(* Logix 5000 project; controller _GigaDiscovery vendor 1 type 14 code 244 rev 35.11; software revision 35.03; part 13 of 23 *)
(* tags used below, declared in another part *)
   OS : DINT;
   Timer : TIMER[60];
   CCW_OS_Direction_1 : BOOL;
   CCW_OS_Direction_2 : BOOL;
   CROUT_Air_Compressor : UDT_CROUT;   // Compressor Command -Q18101E
   CW_OS_Direction_1 : BOOL;
   CW_OS_Direction_2 : BOOL;
   DC_Field_Pylon_Motors : UDT_CROUT;   // DC Field Pylon Motors Contactor -Q10101E -Q10103E
   Emergencies_CL0 : DINT[8];
   Emergencies_CL1 : DINT[14];
   Gate_Entry_Unlock_Selector : BOOL;   // -S30701F
   Gate_Exit_Unlock_Selector : BOOL;   // -S30705F
   Gate_Operator_Unlock_Selector : BOOL;   // -S30707F
   Gondola_Decc_timer_Start : BOOL;
   Gondola_Direction_CW_1 : BOOL;   // 0 > CCW 1 > CW
   Gondola_Direction_CW_2 : BOOL;   // 0 > CCW 1 > CW
   Gondola_Drive_Enable : UDT_CROUT;   // Gondola Drive Ch1-Ch2 Start Enable Contactors -Q16105E -Q16107E
   I_Fbk_Platform_Main_Valve : UDT_DCS;   // Feedback Platform Main Valve -B21902I
   I_GMB_RCC1_Temperature_OK : BOOL;   // +GMB_RCC1 Temperature OK -S40103E
   I_Gondola_Home_Position_Sensor_1 : UDT_DCM;   // Home Sensor Speed Check -B40002I
   I_Gondola_Home_Position_Sensor_2 : UDT_DCM;   // Home Sensor Speed Check -B40007I
   I_OCC2_Disable : UDT_DCM;   // OCC 2 CONTROL DISABLE Page 310
   I_Platform_Closed : UDT_DCM;   // Platform Closed RFID Series -B22501J... -B22807J -B22801B
   I_Platform_Line_Min_Pressure_Switch : BOOL;   // Platform Line Minimum Pressure Switch -S21511B
   I_Platform_Line_Unlock_Pressure_Switch : BOOL;   // Unlock Platform Line Pressure Switch -S22006B
   I_Platform_Opened : UDT_DCM;   // Platform Opened RFID Series -Q23801J -Q23807J
   I_Platform_Pressure_on_Close_Circuit : BOOL;   // Platform Maximum Closing Pressure -S21510B
   I_Pylon_Home_Ch1 : UDT_DCM;   // Home position Pylon Ch1 -B26002I
   I_Pylon_Home_Ch2 : UDT_DCM;   // Home position Pylon Ch2 -B26007I
   I_Pylon_Overlimit_Right : UDT_DCS;   // Pylon Overlimit Switchs -A26510I
   I_RCC_GSA_Temperature_OK : BOOL;   // +RCC_GSA Temperature OK -S50110G
   I_RCC_GSB_Temperature_OK : BOOL;   // +RCC_GSB Temperature OK -S52110G
   I_RCC_GSC_Temperature_OK : BOOL;   // +RCC_GSC Temperature OK -S54110G
   I_RCC_GSD_Temperature_OK : BOOL;   // +RCC_GSD Temperature OK -S56110G
   I_RCC_GSE_Temperature_OK : BOOL;   // +RCC_GSE Temperature OK -S58110G
   I_RCC_GSF_Temperature_OK : BOOL;   // +RCC_GSF Temperature OK -S60110G
   I_RCC_GSG_Temperature_OK : BOOL;   // +RCC_GSG Temperature OK -S62110G
   I_RCC_GSH_Temperature_OK : BOOL;   // +RCC_GSH Temperature OK -S64110G
   Max_Gondola_Speed_RPM : REAL;
   Max_Gondola_Speed_RPS : REAL;
   No_Sfty : Std_to_Sfty;
   No_Sfty_Gondola_SpdFeedback_ABS : DINT;
   O_Pilots_Valve_Platform : BOOL;
   O_Platform_Main_Valve : BOOL;   // Valvola principale piattaforma B21902I
   O_Platform_MainValve : UDT_CROUT;   // Platform main valve B21902I
   ONP : DINT;   // Optional Not Present
   Overspeed_Threshold_millisec : DINT;
   Overspeed_Threshold_sec : REAL;
   Platform_Close_Cycle : Sequencer;
   Platform_Closing_Cycle_Alarms_Ok : BOOL;
   Platform_Fbk_Valv_Open : BOOL;   // Platform Open Main Valve Limit Switch -B21905I
   Platform_Open_Cycle : Sequencer;
   Power_On_Delay : BOOL;
   ProofTest_Req : BOOL;
   Pylon_Brake_Motor : UDT_CROUT;   // Pylon Brake command -Q10801E
   Pylon_Overspeed_Max_Th : DINT;
   Pylon_Overspeed_min_Th : DINT;
   Pylon_Overspeed_Sensors : DCA_INPUT;
   Pylon_Speed : DINT;
   Reset_Pulse : BOOL;
   RESTRAINTS_Closed : BOOL;   // All RESTRAINTS Closed
   Restraints_Cycle : Sequencer;
   RESTRAINTS_Left_Press_Switch_Series : BOOL;
   RESTRAINTS_No_Alarms : BOOL;
   RESTRAINTS_Right_Press_Switch_Series : BOOL;
   RESTRAINTS_Sector : LapBars_Sector[9];
   Revolution_time_1 : DINT;
   Revolution_time_2 : DINT;
   Speed_at_Minute : REAL;
   Speed_at_Second : REAL;
   Start_Stop_Cycle : Sequencer;
   Stop_Request : BOOL;
   Timer_Overspeed_reset_1 : BOOL;   // senor 1 Revolution time reset
   Timer_Overspeed_reset_2 : BOOL;   // senor 2
   Valve_Proof_Test_Cycle : Sequencer;
(* S_Alarms, continued *)

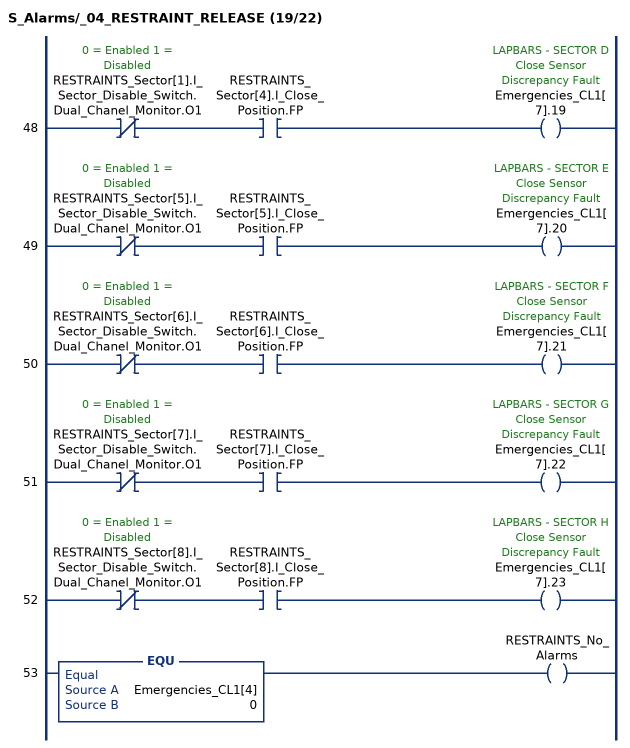
   [picture p233: S_Alarms/_04_RESTRAINT_RELEASE rungs 48-53]
   48: XIO(RESTRAINTS_Sector[1].I_Sector_Disable_Switch.Dual_Chanel_Monitor.O1)XIC(RESTRAINTS_Sector[4].I_Close_Position.FP)OTE(Emergencies_CL1[7].19);
   49: XIO(RESTRAINTS_Sector[5].I_Sector_Disable_Switch.Dual_Chanel_Monitor.O1)XIC(RESTRAINTS_Sector[5].I_Close_Position.FP)OTE(Emergencies_CL1[7].20);
   50: XIO(RESTRAINTS_Sector[6].I_Sector_Disable_Switch.Dual_Chanel_Monitor.O1)XIC(RESTRAINTS_Sector[6].I_Close_Position.FP)OTE(Emergencies_CL1[7].21);
   51: XIO(RESTRAINTS_Sector[7].I_Sector_Disable_Switch.Dual_Chanel_Monitor.O1)XIC(RESTRAINTS_Sector[7].I_Close_Position.FP)OTE(Emergencies_CL1[7].22);
   52: XIO(RESTRAINTS_Sector[8].I_Sector_Disable_Switch.Dual_Chanel_Monitor.O1)XIC(RESTRAINTS_Sector[8].I_Close_Position.FP)OTE(Emergencies_CL1[7].23);
   53: EQU(Emergencies_CL1[4],0)OTE(RESTRAINTS_No_Alarms);
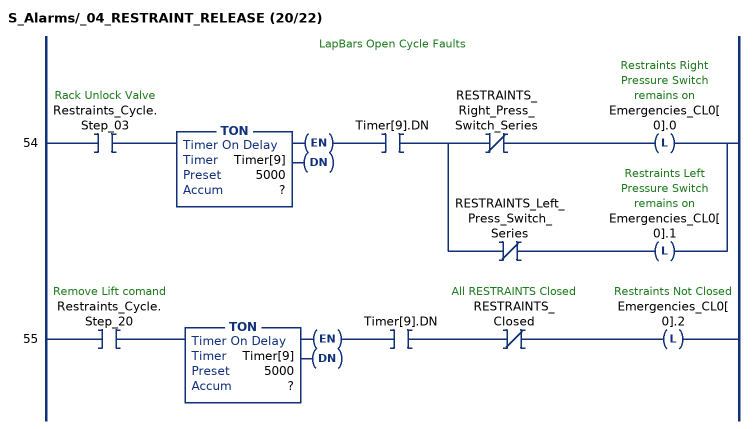
   // LapBars Open Cycle Faults
   54: XIC(Restraints_Cycle.Step_03)TON(Timer[9],?,?)XIC(Timer[9].DN)[XIO(RESTRAINTS_Right_Press_Switch_Series) OTL(Emergencies_CL0[0].0) ,XIO(RESTRAINTS_Left_Press_Switch_Series) OTL(Emergencies_CL0[0].1) ];
   55: XIC(Restraints_Cycle.Step_20)TON(Timer[9],?,?)XIC(Timer[9].DN)XIO(RESTRAINTS_Closed)OTL(Emergencies_CL0[0].2);
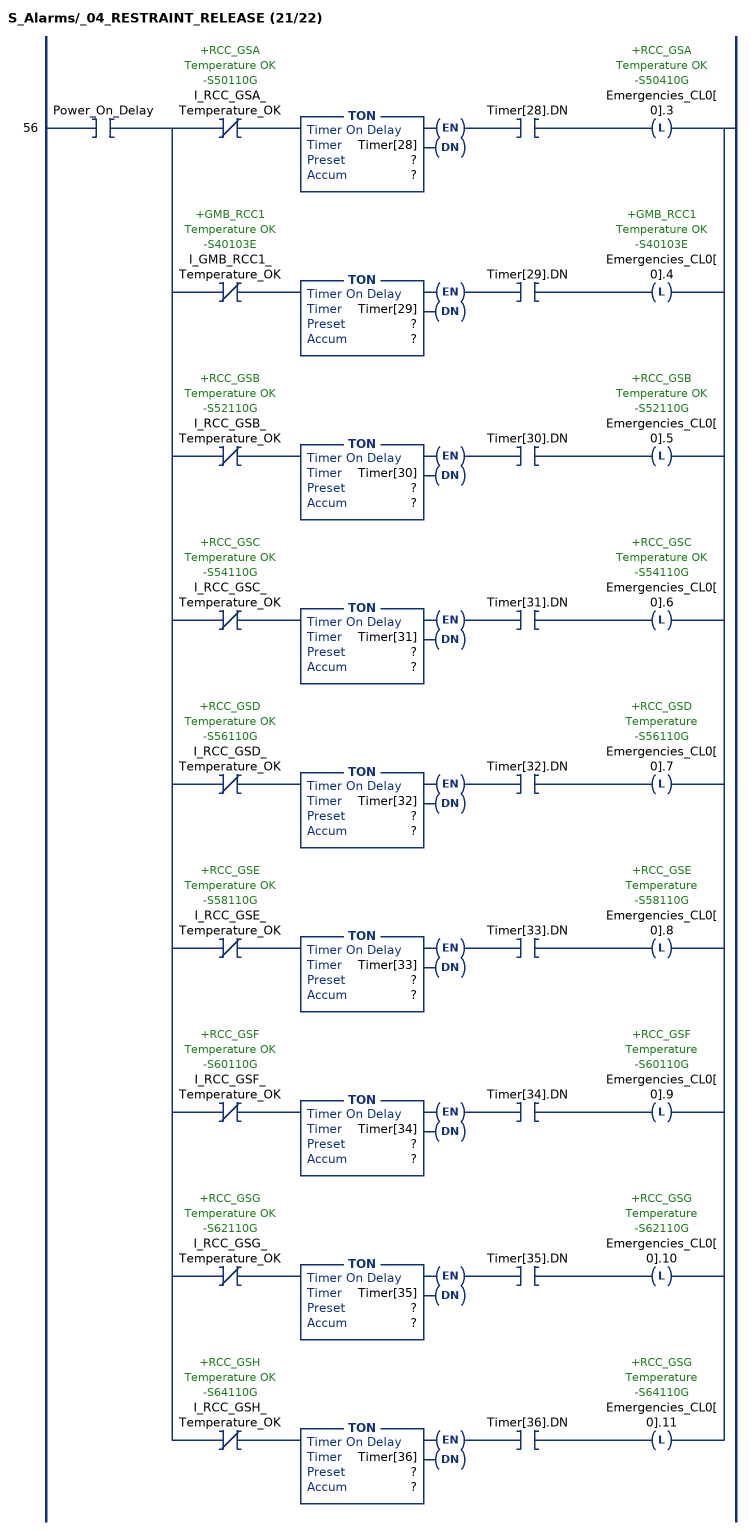
   56: XIC(Power_On_Delay)[XIO(I_RCC_GSA_Temperature_OK) TON(Timer[28],?,?) XIC(Timer[28].DN) OTL(Emergencies_CL0[0].3) ,XIO(I_GMB_RCC1_Temperature_OK) TON(Timer[29],?,?) XIC(Timer[29].DN) OTL(Emergencies_CL0[0].4) ,XIO(I_RCC_GSB_Temperature_OK) TON(Timer[30],?,?) XIC(Timer[30].DN) OTL(Emergencies_CL0[0].5) ,XIO(I_RCC_GSC_Temperature_OK) TON(Timer[31],?,?) XIC(Timer[31].DN) OTL(Emergencies_CL0[0].6) ,XIO(I_RCC_GSD_Temperature_OK) TON(Timer[32],?,?) XIC(Timer[32].DN) OTL(Emergencies_CL0[0].7) ,XIO(I_RCC_GSE_Temperature_OK) TON(Timer[33],?,?) XIC(Timer[33].DN) OTL(Emergencies_CL0[0].8) ,XIO(I_RCC_GSF_Temperature_OK) TON(Timer[34],?,?) XIC(Timer[34].DN) OTL(Emergencies_CL0[0].9) ,XIO(I_RCC_GSG_Temperature_OK) TON(Timer[35],?,?) XIC(Timer[35].DN) OTL(Emergencies_CL0[0].10) ,XIO(I_RCC_GSH_Temperature_OK) TON(Timer[36],?,?) XIC(Timer[36].DN) OTL(Emergencies_CL0[0].11) ];
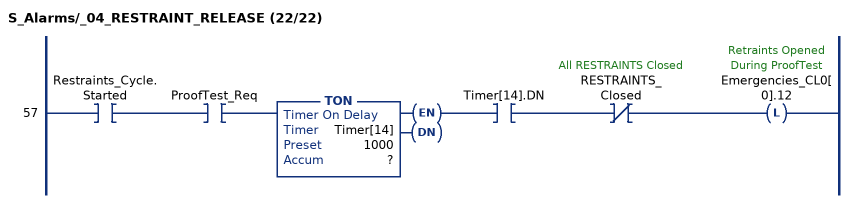
   57: XIC(Restraints_Cycle.Started)XIC(ProofTest_Req)TON(Timer[14],?,?)XIC(Timer[14].DN)XIO(RESTRAINTS_Closed)OTL(Emergencies_CL0[0].12);
END_ROUTINE

ROUTINE _05_Platform   (* ladder *)
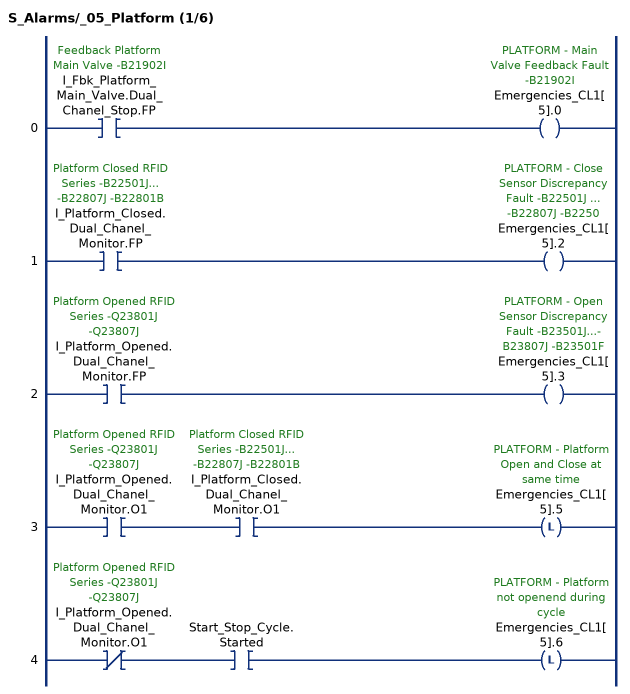
   0: XIC(I_Fbk_Platform_Main_Valve.Dual_Chanel_Stop.FP)OTE(Emergencies_CL1[5].0);
   1: XIC(I_Platform_Closed.Dual_Chanel_Monitor.FP)OTE(Emergencies_CL1[5].2);
   2: XIC(I_Platform_Opened.Dual_Chanel_Monitor.FP)OTE(Emergencies_CL1[5].3);
   3: XIC(I_Platform_Opened.Dual_Chanel_Monitor.O1)XIC(I_Platform_Closed.Dual_Chanel_Monitor.O1)OTL(Emergencies_CL1[5].5);
   4: XIO(I_Platform_Opened.Dual_Chanel_Monitor.O1)XIC(Start_Stop_Cycle.Started)OTL(Emergencies_CL1[5].6);
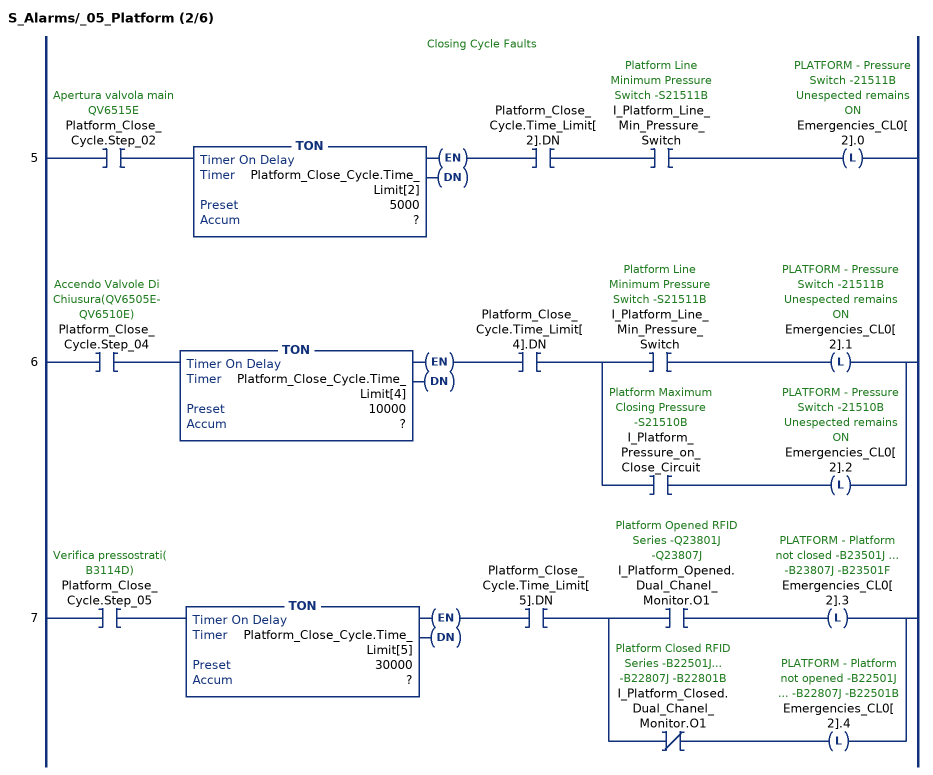
   // Closing Cycle Faults
   5: XIC(Platform_Close_Cycle.Step_02)TON(Platform_Close_Cycle.Time_Limit[2],?,?)XIC(Platform_Close_Cycle.Time_Limit[2].DN)XIC(I_Platform_Line_Min_Pressure_Switch)OTL(Emergencies_CL0[2].0);
   6: XIC(Platform_Close_Cycle.Step_04)TON(Platform_Close_Cycle.Time_Limit[4],?,?)XIC(Platform_Close_Cycle.Time_Limit[4].DN)[XIC(I_Platform_Line_Min_Pressure_Switch) OTL(Emergencies_CL0[2].1) ,XIC(I_Platform_Pressure_on_Close_Circuit) OTL(Emergencies_CL0[2].2) ];
   7: XIC(Platform_Close_Cycle.Step_05)TON(Platform_Close_Cycle.Time_Limit[5],?,?)XIC(Platform_Close_Cycle.Time_Limit[5].DN)[XIC(I_Platform_Opened.Dual_Chanel_Monitor.O1) OTL(Emergencies_CL0[2].3) ,XIO(I_Platform_Closed.Dual_Chanel_Monitor.O1) OTL(Emergencies_CL0[2].4) ];
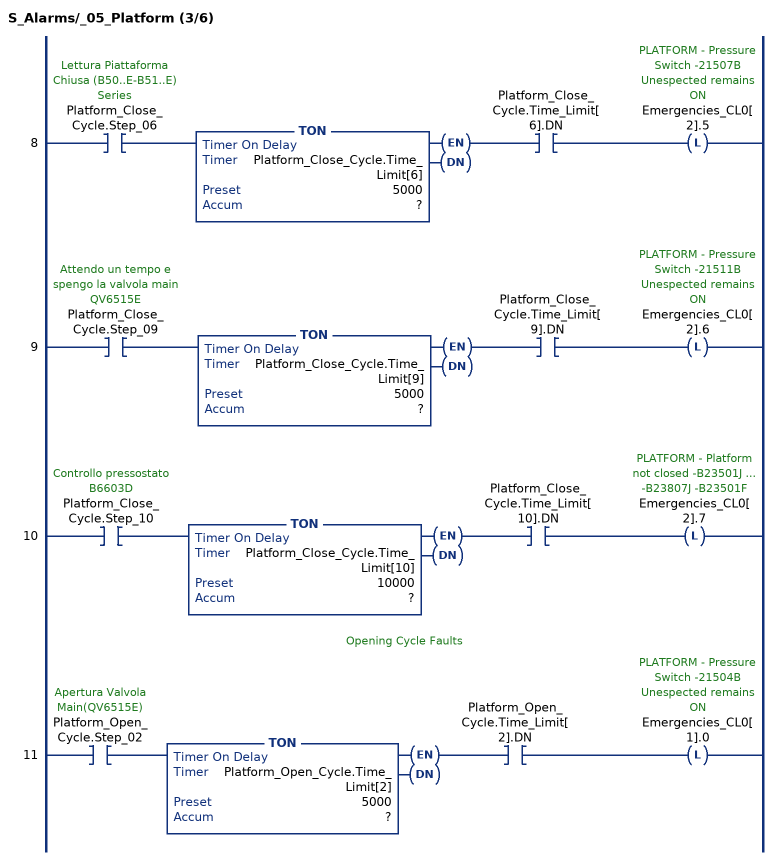
   8: XIC(Platform_Close_Cycle.Step_06)TON(Platform_Close_Cycle.Time_Limit[6],?,?)XIC(Platform_Close_Cycle.Time_Limit[6].DN)OTL(Emergencies_CL0[2].5);
   9: XIC(Platform_Close_Cycle.Step_09)TON(Platform_Close_Cycle.Time_Limit[9],?,?)XIC(Platform_Close_Cycle.Time_Limit[9].DN)OTL(Emergencies_CL0[2].6);
   10: XIC(Platform_Close_Cycle.Step_10)TON(Platform_Close_Cycle.Time_Limit[10],?,?)XIC(Platform_Close_Cycle.Time_Limit[10].DN)OTL(Emergencies_CL0[2].7);
   // Opening Cycle Faults
   11: XIC(Platform_Open_Cycle.Step_02)TON(Platform_Open_Cycle.Time_Limit[2],?,?)XIC(Platform_Open_Cycle.Time_Limit[2].DN)OTL(Emergencies_CL0[1].0);
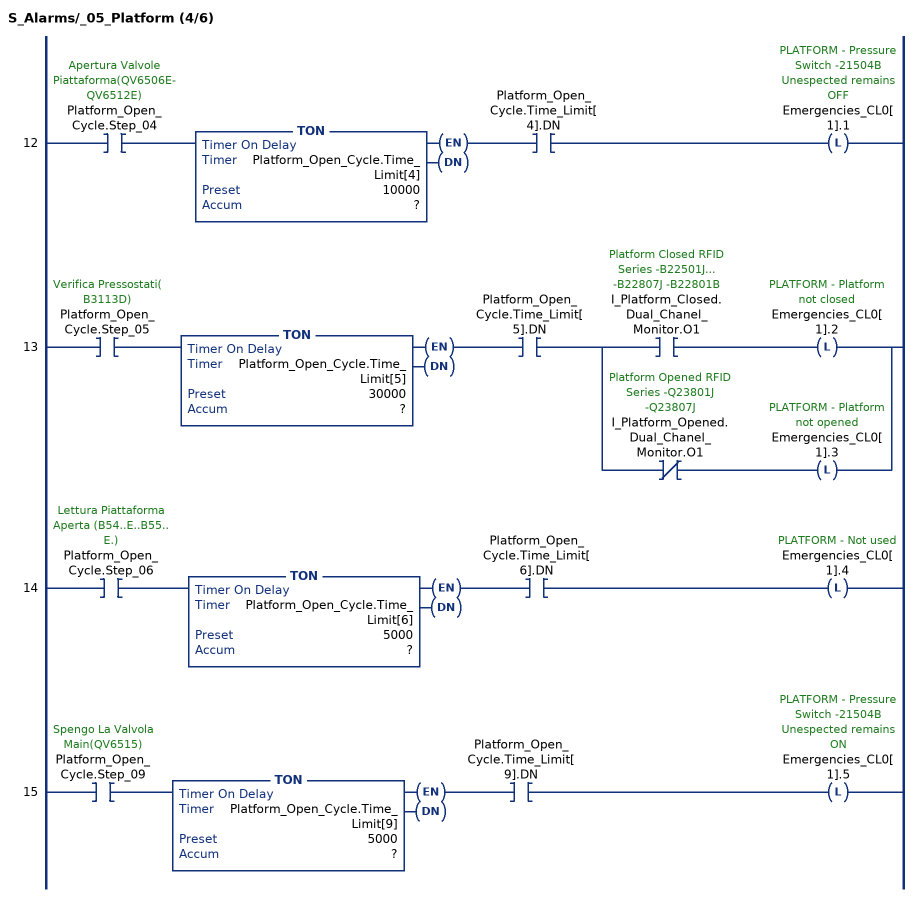
   12: XIC(Platform_Open_Cycle.Step_04)TON(Platform_Open_Cycle.Time_Limit[4],?,?)XIC(Platform_Open_Cycle.Time_Limit[4].DN)OTL(Emergencies_CL0[1].1);
   13: XIC(Platform_Open_Cycle.Step_05)TON(Platform_Open_Cycle.Time_Limit[5],?,?)XIC(Platform_Open_Cycle.Time_Limit[5].DN)[XIC(I_Platform_Closed.Dual_Chanel_Monitor.O1) OTL(Emergencies_CL0[1].2) ,XIO(I_Platform_Opened.Dual_Chanel_Monitor.O1) OTL(Emergencies_CL0[1].3) ];
   14: XIC(Platform_Open_Cycle.Step_06)TON(Platform_Open_Cycle.Time_Limit[6],?,?)XIC(Platform_Open_Cycle.Time_Limit[6].DN)OTL(Emergencies_CL0[1].4);
   15: XIC(Platform_Open_Cycle.Step_09)TON(Platform_Open_Cycle.Time_Limit[9],?,?)XIC(Platform_Open_Cycle.Time_Limit[9].DN)OTL(Emergencies_CL0[1].5);
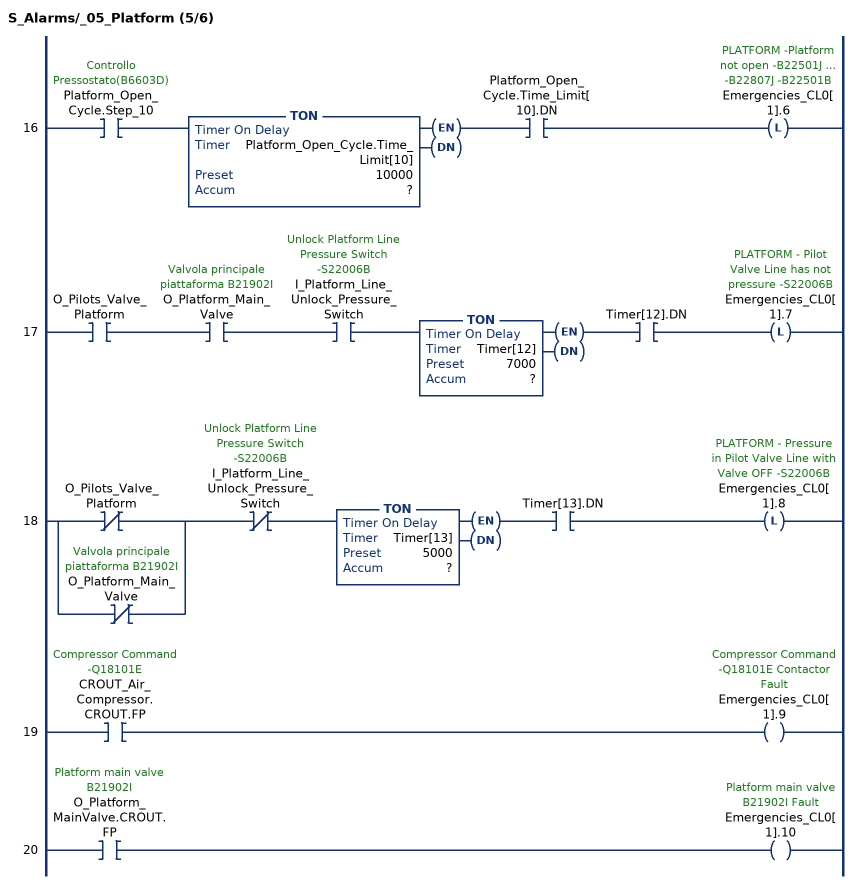
   16: XIC(Platform_Open_Cycle.Step_10)TON(Platform_Open_Cycle.Time_Limit[10],?,?)XIC(Platform_Open_Cycle.Time_Limit[10].DN)OTL(Emergencies_CL0[1].6);
   17: XIC(O_Pilots_Valve_Platform)XIC(O_Platform_Main_Valve)XIC(I_Platform_Line_Unlock_Pressure_Switch)TON(Timer[12],?,?)XIC(Timer[12].DN)OTL(Emergencies_CL0[1].7);
   18: [XIO(O_Pilots_Valve_Platform) ,XIO(O_Platform_Main_Valve) ]XIO(I_Platform_Line_Unlock_Pressure_Switch)TON(Timer[13],?,?)XIC(Timer[13].DN)OTL(Emergencies_CL0[1].8);
   19: XIC(CROUT_Air_Compressor.CROUT.FP)OTE(Emergencies_CL0[1].9);
   20: XIC(O_Platform_MainValve.CROUT.FP)OTE(Emergencies_CL0[1].10);
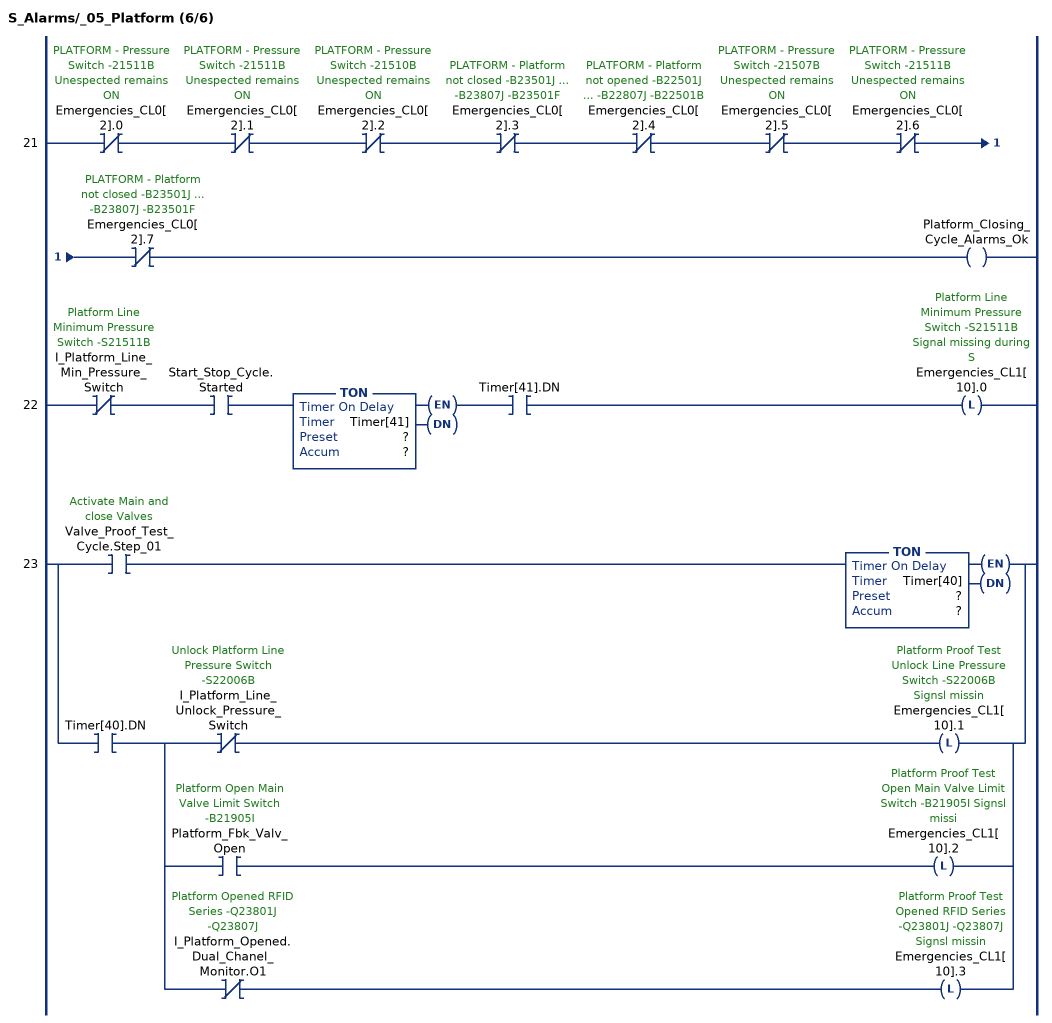
   21: XIO(Emergencies_CL0[2].0)XIO(Emergencies_CL0[2].1)XIO(Emergencies_CL0[2].2)XIO(Emergencies_CL0[2].3)XIO(Emergencies_CL0[2].4)XIO(Emergencies_CL0[2].5)XIO(Emergencies_CL0[2].6)XIO(Emergencies_CL0[2].7)OTE(Platform_Closing_Cycle_Alarms_Ok);
   22: XIO(I_Platform_Line_Min_Pressure_Switch)XIC(Start_Stop_Cycle.Started)TON(Timer[41],?,?)XIC(Timer[41].DN)OTL(Emergencies_CL1[10].0);
   23: [XIC(Valve_Proof_Test_Cycle.Step_01) TON(Timer[40],?,?) ,XIC(Timer[40].DN) [XIO(I_Platform_Line_Unlock_Pressure_Switch) OTL(Emergencies_CL1[10].1) ,XIC(Platform_Fbk_Valv_Open) OTL(Emergencies_CL1[10].2) ,XIO(I_Platform_Opened.Dual_Chanel_Monitor.O1) OTL(Emergencies_CL1[10].3) ] ];
END_ROUTINE

ROUTINE _06_Pylon_Gondola   (* ladder *)
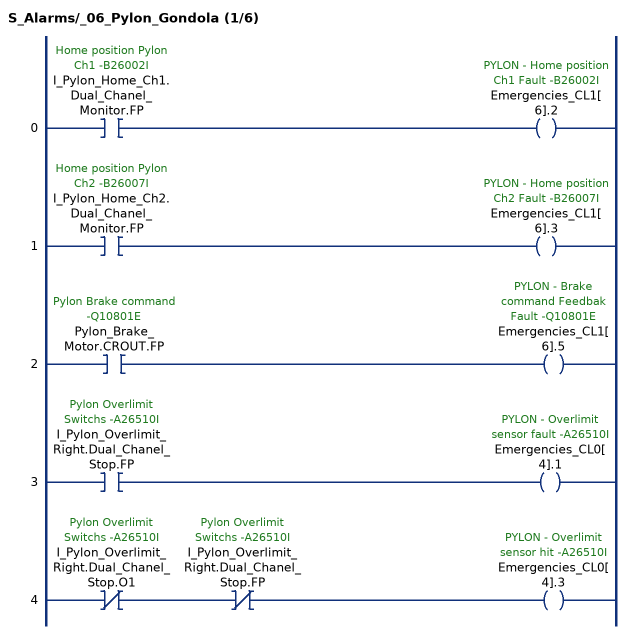
   0: XIC(I_Pylon_Home_Ch1.Dual_Chanel_Monitor.FP)OTE(Emergencies_CL1[6].2);
   1: XIC(I_Pylon_Home_Ch2.Dual_Chanel_Monitor.FP)OTE(Emergencies_CL1[6].3);
   2: XIC(Pylon_Brake_Motor.CROUT.FP)OTE(Emergencies_CL1[6].5);
   3: XIC(I_Pylon_Overlimit_Right.Dual_Chanel_Stop.FP)OTE(Emergencies_CL0[4].1);
   4: XIO(I_Pylon_Overlimit_Right.Dual_Chanel_Stop.O1)XIO(I_Pylon_Overlimit_Right.Dual_Chanel_Stop.FP)OTE(Emergencies_CL0[4].3);
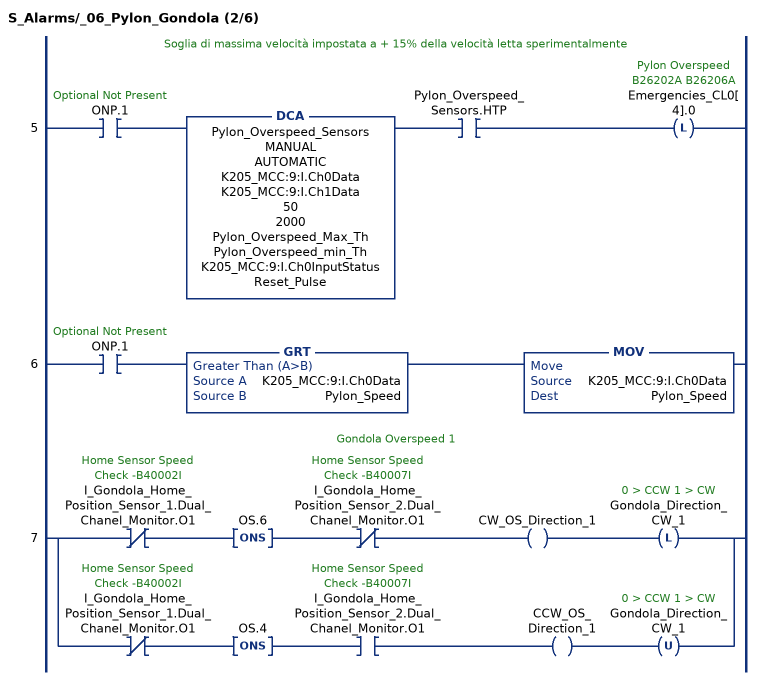
   // Soglia di massima velocità impostata a + 15% della velocità letta sperimentalmente
   5: XIC(ONP.1)DCA(Pylon_Overspeed_Sensors,MANUAL,AUTOMATIC,K205_MCC:9:I.Ch0Data,K205_MCC:9:I.Ch1Data,50,2000,Pylon_Overspeed_Max_Th,Pylon_Overspeed_min_Th,K205_MCC:9:I.Ch0InputStatus,Reset_Pulse)XIC(Pylon_Overspeed_Sensors.HTP)OTL(Emergencies_CL0[4].0);
   6: XIC(ONP.1)GRT(K205_MCC:9:I.Ch0Data,Pylon_Speed)MOV(K205_MCC:9:I.Ch0Data,Pylon_Speed);
   // Gondola Overspeed 1
   7: [XIO(I_Gondola_Home_Position_Sensor_1.Dual_Chanel_Monitor.O1) ONS(OS.6) XIO(I_Gondola_Home_Position_Sensor_2.Dual_Chanel_Monitor.O1) OTE(CW_OS_Direction_1) OTL(Gondola_Direction_CW_1) ,XIO(I_Gondola_Home_Position_Sensor_1.Dual_Chanel_Monitor.O1) ONS(OS.4) XIC(I_Gondola_Home_Position_Sensor_2.Dual_Chanel_Monitor.O1) OTE(CCW_OS_Direction_1) OTU(Gondola_Direction_CW_1) ];
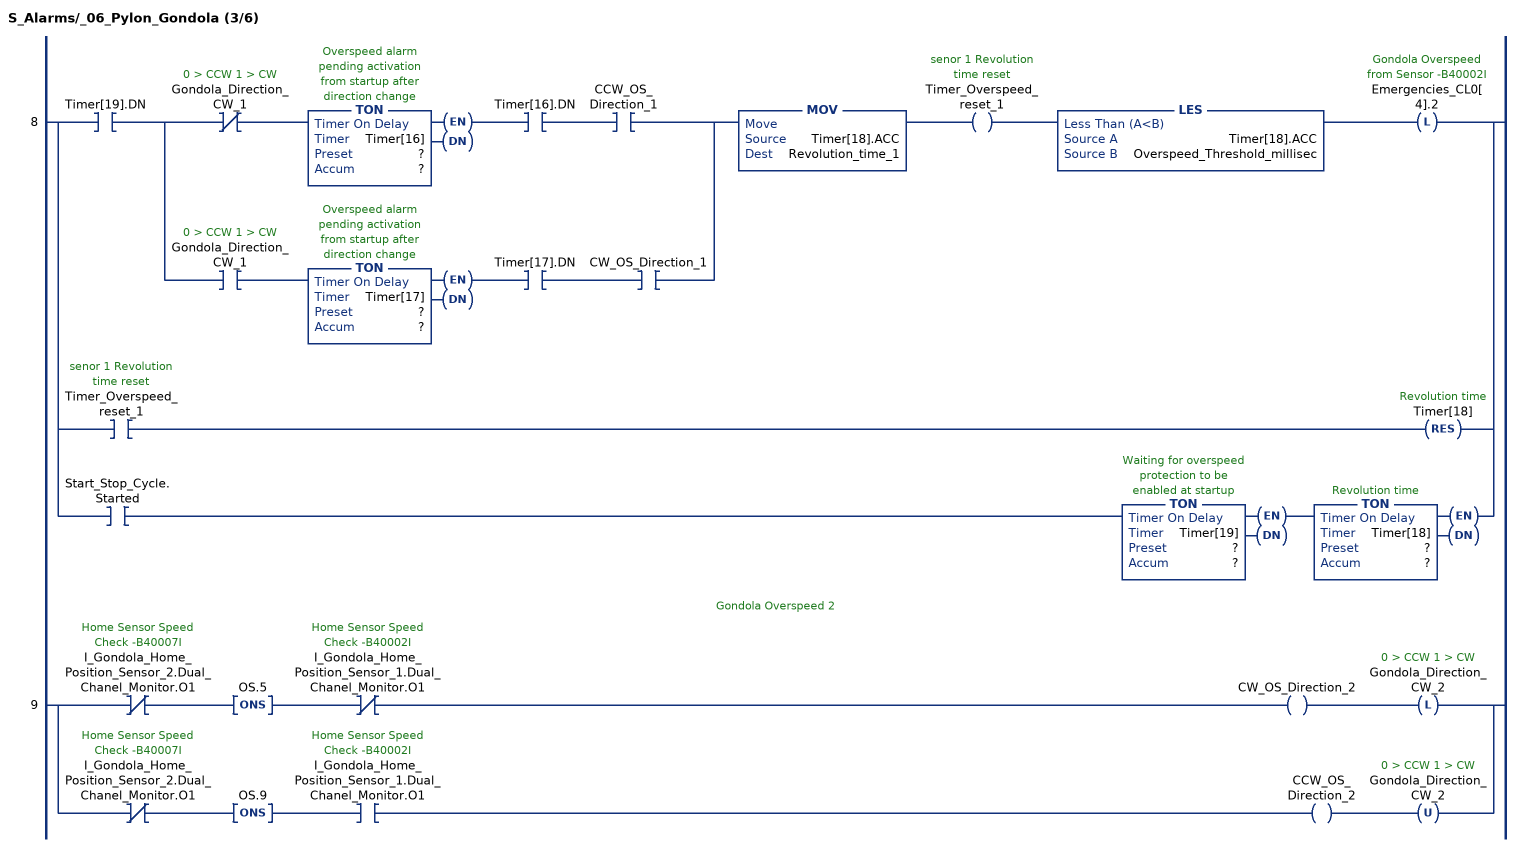
   8: [XIC(Timer[19].DN) [XIO(Gondola_Direction_CW_1) TON(Timer[16],?,?) XIC(Timer[16].DN) XIC(CCW_OS_Direction_1) ,XIC(Gondola_Direction_CW_1) TON(Timer[17],?,?) XIC(Timer[17].DN) XIC(CW_OS_Direction_1) ] MOV(Timer[18].ACC,Revolution_time_1) OTE(Timer_Overspeed_reset_1) LES(Timer[18].ACC,Overspeed_Threshold_millisec) OTL(Emergencies_CL0[4].2) ,XIC(Timer_Overspeed_reset_1) RES(Timer[18]) ,XIC(Start_Stop_Cycle.Started) TON(Timer[19],?,?) TON(Timer[18],?,?) ];
   // Gondola Overspeed 2
   9: [XIO(I_Gondola_Home_Position_Sensor_2.Dual_Chanel_Monitor.O1) ONS(OS.5) XIO(I_Gondola_Home_Position_Sensor_1.Dual_Chanel_Monitor.O1) OTE(CW_OS_Direction_2) OTL(Gondola_Direction_CW_2) ,XIO(I_Gondola_Home_Position_Sensor_2.Dual_Chanel_Monitor.O1) ONS(OS.9) XIC(I_Gondola_Home_Position_Sensor_1.Dual_Chanel_Monitor.O1) OTE(CCW_OS_Direction_2) OTU(Gondola_Direction_CW_2) ];
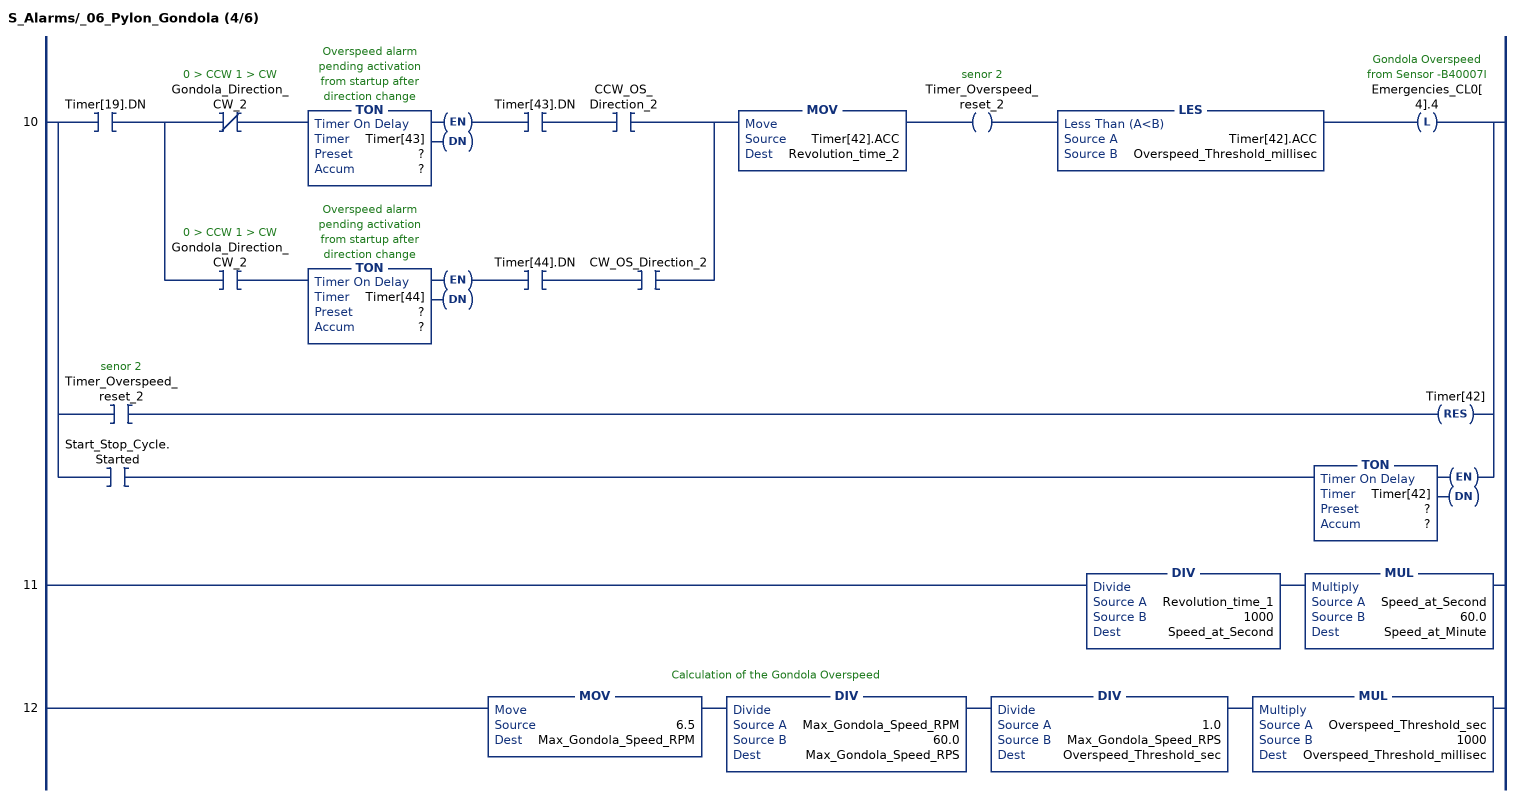
   10: [XIC(Timer[19].DN) [XIO(Gondola_Direction_CW_2) TON(Timer[43],?,?) XIC(Timer[43].DN) XIC(CCW_OS_Direction_2) ,XIC(Gondola_Direction_CW_2) TON(Timer[44],?,?) XIC(Timer[44].DN) XIC(CW_OS_Direction_2) ] MOV(Timer[42].ACC,Revolution_time_2) OTE(Timer_Overspeed_reset_2) LES(Timer[42].ACC,Overspeed_Threshold_millisec) OTL(Emergencies_CL0[4].4) ,XIC(Timer_Overspeed_reset_2) RES(Timer[42]) ,XIC(Start_Stop_Cycle.Started) TON(Timer[42],?,?) ];
   11: DIV(Revolution_time_1,1000,Speed_at_Second)MUL(Speed_at_Second,60.0,Speed_at_Minute);
   // Calculation of the Gondola Overspeed
   12: MOV(6.5,Max_Gondola_Speed_RPM)DIV(Max_Gondola_Speed_RPM,60.0,Max_Gondola_Speed_RPS)DIV(1.0,Max_Gondola_Speed_RPS,Overspeed_Threshold_sec)MUL(Overspeed_Threshold_sec,1000,Overspeed_Threshold_millisec);
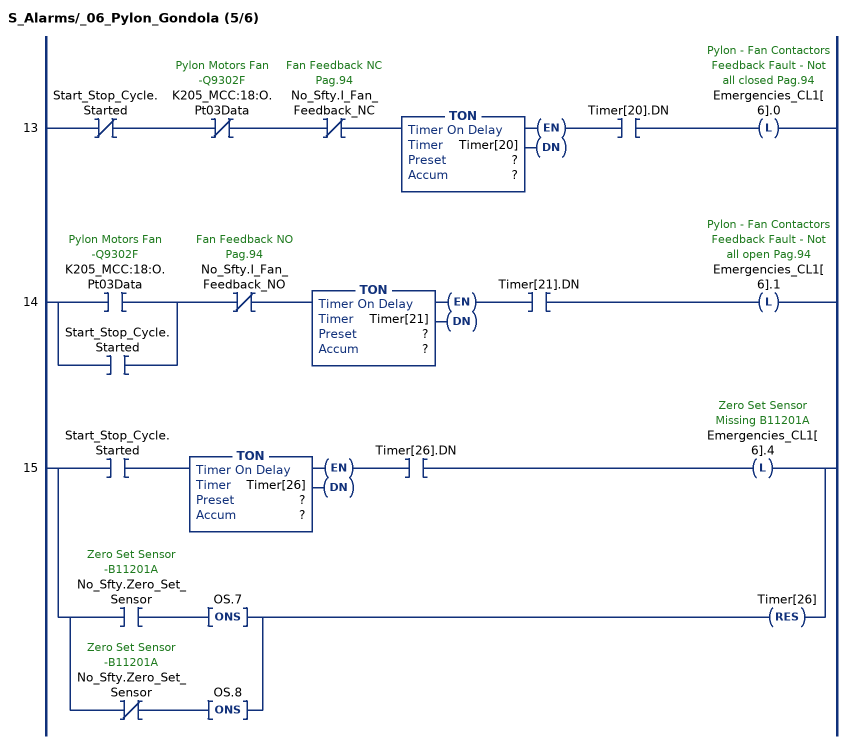
   13: XIO(Start_Stop_Cycle.Started)XIO(K205_MCC:18:O.Pt03Data)XIO(No_Sfty.I_Fan_Feedback_NC)TON(Timer[20],?,?)XIC(Timer[20].DN)OTL(Emergencies_CL1[6].0);
   14: [XIC(K205_MCC:18:O.Pt03Data) ,XIC(Start_Stop_Cycle.Started) ]XIO(No_Sfty.I_Fan_Feedback_NO)TON(Timer[21],?,?)XIC(Timer[21].DN)OTL(Emergencies_CL1[6].1);
   15: [XIC(Start_Stop_Cycle.Started) TON(Timer[26],?,?) XIC(Timer[26].DN) OTL(Emergencies_CL1[6].4) ,[XIC(No_Sfty.Zero_Set_Sensor) ONS(OS.7) ,XIO(No_Sfty.Zero_Set_Sensor) ONS(OS.8) ] RES(Timer[26]) ];
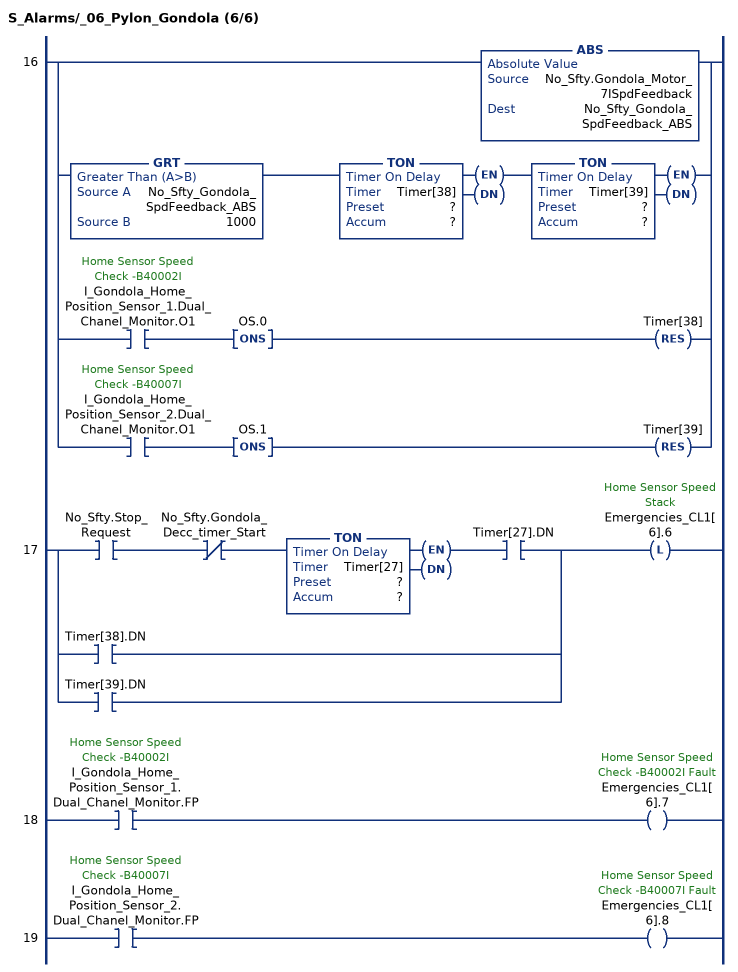
   16: [ABS(No_Sfty.Gondola_Motor_7ISpdFeedback,No_Sfty_Gondola_SpdFeedback_ABS) ,GRT(No_Sfty_Gondola_SpdFeedback_ABS,1000) TON(Timer[38],?,?) TON(Timer[39],?,?) ,XIC(I_Gondola_Home_Position_Sensor_1.Dual_Chanel_Monitor.O1) ONS(OS.0) RES(Timer[38]) ,XIC(I_Gondola_Home_Position_Sensor_2.Dual_Chanel_Monitor.O1) ONS(OS.1) RES(Timer[39]) ];
   17: [XIC(No_Sfty.Stop_Request) XIO(No_Sfty.Gondola_Decc_timer_Start) TON(Timer[27],?,?) XIC(Timer[27].DN) ,XIC(Timer[38].DN) ,XIC(Timer[39].DN) ]OTL(Emergencies_CL1[6].6);
   18: XIC(I_Gondola_Home_Position_Sensor_1.Dual_Chanel_Monitor.FP)OTE(Emergencies_CL1[6].7);
   19: XIC(I_Gondola_Home_Position_Sensor_2.Dual_Chanel_Monitor.FP)OTE(Emergencies_CL1[6].8);
END_ROUTINE

ROUTINE _07_Auto_Cycle   (* ladder *)
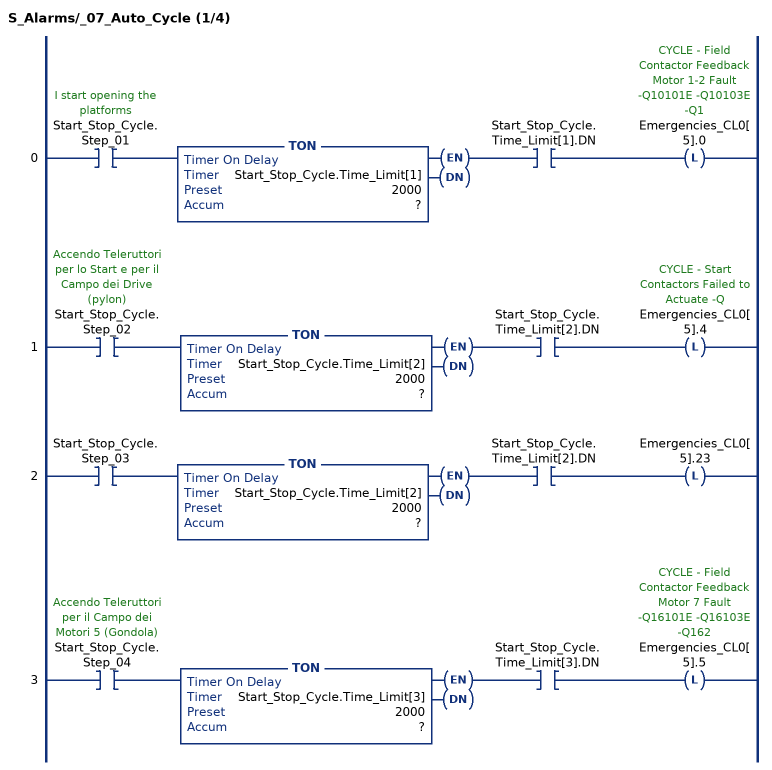
   0: XIC(Start_Stop_Cycle.Step_01)TON(Start_Stop_Cycle.Time_Limit[1],?,?)XIC(Start_Stop_Cycle.Time_Limit[1].DN)OTL(Emergencies_CL0[5].0);
   1: XIC(Start_Stop_Cycle.Step_02)TON(Start_Stop_Cycle.Time_Limit[2],?,?)XIC(Start_Stop_Cycle.Time_Limit[2].DN)OTL(Emergencies_CL0[5].4);
   2: XIC(Start_Stop_Cycle.Step_03)TON(Start_Stop_Cycle.Time_Limit[2],?,?)XIC(Start_Stop_Cycle.Time_Limit[2].DN)OTL(Emergencies_CL0[5].23);
   3: XIC(Start_Stop_Cycle.Step_04)TON(Start_Stop_Cycle.Time_Limit[3],?,?)XIC(Start_Stop_Cycle.Time_Limit[3].DN)OTL(Emergencies_CL0[5].5);
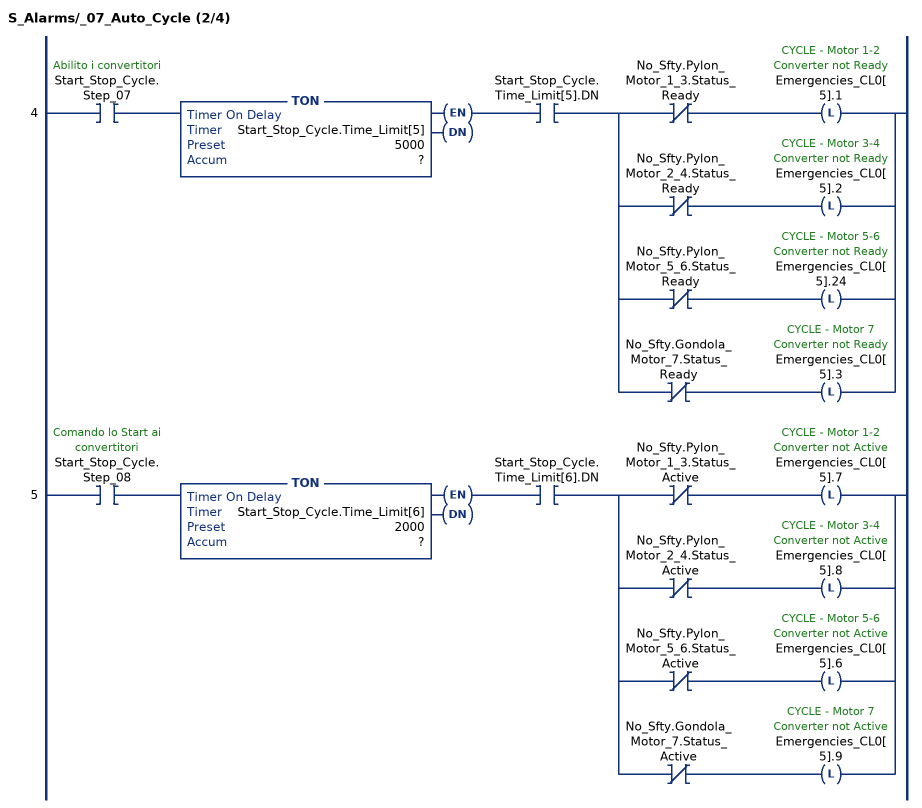
   4: XIC(Start_Stop_Cycle.Step_07)TON(Start_Stop_Cycle.Time_Limit[5],?,?)XIC(Start_Stop_Cycle.Time_Limit[5].DN)[XIO(No_Sfty.Pylon_Motor_1_3.Status_Ready) OTL(Emergencies_CL0[5].1) ,XIO(No_Sfty.Pylon_Motor_2_4.Status_Ready) OTL(Emergencies_CL0[5].2) ,XIO(No_Sfty.Pylon_Motor_5_6.Status_Ready) OTL(Emergencies_CL0[5].24) ,XIO(No_Sfty.Gondola_Motor_7.Status_Ready) OTL(Emergencies_CL0[5].3) ];
   5: XIC(Start_Stop_Cycle.Step_08)TON(Start_Stop_Cycle.Time_Limit[6],?,?)XIC(Start_Stop_Cycle.Time_Limit[6].DN)[XIO(No_Sfty.Pylon_Motor_1_3.Status_Active) OTL(Emergencies_CL0[5].7) ,XIO(No_Sfty.Pylon_Motor_2_4.Status_Active) OTL(Emergencies_CL0[5].8) ,XIO(No_Sfty.Pylon_Motor_5_6.Status_Active) OTL(Emergencies_CL0[5].6) ,XIO(No_Sfty.Gondola_Motor_7.Status_Active) OTL(Emergencies_CL0[5].9) ];
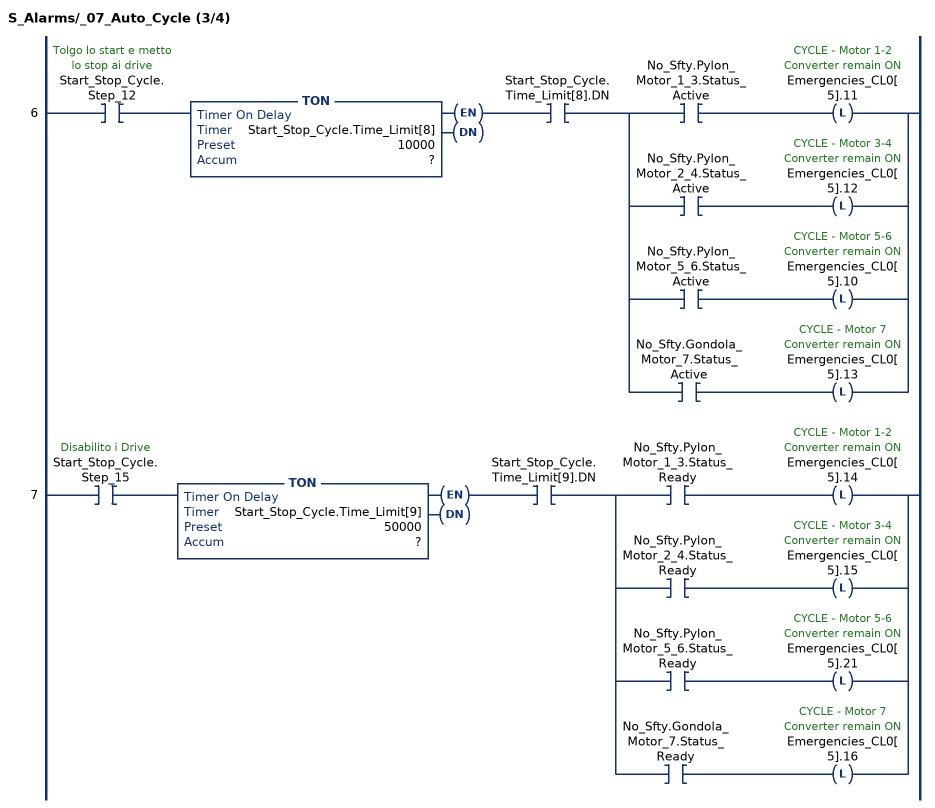
   6: XIC(Start_Stop_Cycle.Step_12)TON(Start_Stop_Cycle.Time_Limit[8],?,?)XIC(Start_Stop_Cycle.Time_Limit[8].DN)[XIC(No_Sfty.Pylon_Motor_1_3.Status_Active) OTL(Emergencies_CL0[5].11) ,XIC(No_Sfty.Pylon_Motor_2_4.Status_Active) OTL(Emergencies_CL0[5].12) ,XIC(No_Sfty.Pylon_Motor_5_6.Status_Active) OTL(Emergencies_CL0[5].10) ,XIC(No_Sfty.Gondola_Motor_7.Status_Active) OTL(Emergencies_CL0[5].13) ];
   7: XIC(Start_Stop_Cycle.Step_15)TON(Start_Stop_Cycle.Time_Limit[9],?,?)XIC(Start_Stop_Cycle.Time_Limit[9].DN)[XIC(No_Sfty.Pylon_Motor_1_3.Status_Ready) OTL(Emergencies_CL0[5].14) ,XIC(No_Sfty.Pylon_Motor_2_4.Status_Ready) OTL(Emergencies_CL0[5].15) ,XIC(No_Sfty.Pylon_Motor_5_6.Status_Ready) OTL(Emergencies_CL0[5].21) ,XIC(No_Sfty.Gondola_Motor_7.Status_Ready) OTL(Emergencies_CL0[5].16) ];
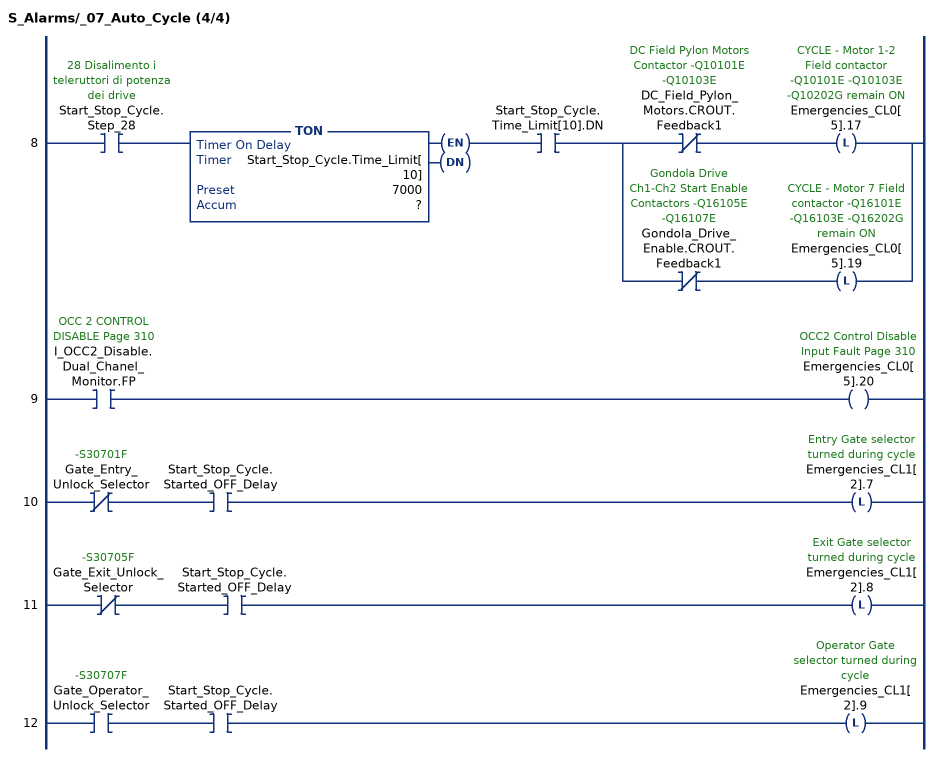
   8: XIC(Start_Stop_Cycle.Step_28)TON(Start_Stop_Cycle.Time_Limit[10],?,?)XIC(Start_Stop_Cycle.Time_Limit[10].DN)[XIO(DC_Field_Pylon_Motors.CROUT.Feedback1) OTL(Emergencies_CL0[5].17) ,XIO(Gondola_Drive_Enable.CROUT.Feedback1) OTL(Emergencies_CL0[5].19) ];
   9: XIC(I_OCC2_Disable.Dual_Chanel_Monitor.FP)OTE(Emergencies_CL0[5].20);
   10: XIO(Gate_Entry_Unlock_Selector)XIC(Start_Stop_Cycle.Started_OFF_Delay)OTL(Emergencies_CL1[2].7);
   11: XIO(Gate_Exit_Unlock_Selector)XIC(Start_Stop_Cycle.Started_OFF_Delay)OTL(Emergencies_CL1[2].8);
   12: XIC(Gate_Operator_Unlock_Selector)XIC(Start_Stop_Cycle.Started_OFF_Delay)OTL(Emergencies_CL1[2].9);
END_ROUTINE
